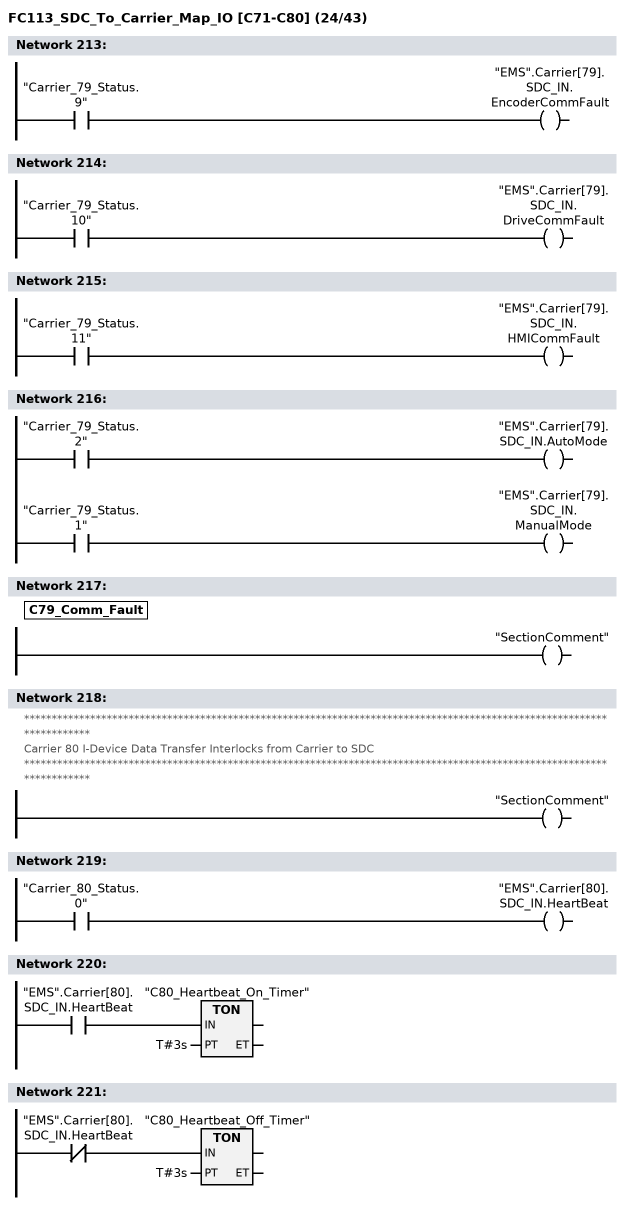
   RUNG wire#powerrail
      Contact( "Carrier_79_Status.9" )
      Coil( "EMS".Carrier[79].SDC_IN.EncoderCommFault )
   END_RUNG
   // the same network as SCL:
   "EMS".Carrier[79].SDC_IN.EncoderCommFault := "Carrier_79_Status.9";
END_REGION

REGION Network 214
   RUNG wire#powerrail
      Contact( "Carrier_79_Status.10" )
      Coil( "EMS".Carrier[79].SDC_IN.DriveCommFault )
   END_RUNG
   // the same network as SCL:
   "EMS".Carrier[79].SDC_IN.DriveCommFault := "Carrier_79_Status.10";
END_REGION

REGION Network 215
   RUNG wire#powerrail
      Contact( "Carrier_79_Status.11" )
      Coil( "EMS".Carrier[79].SDC_IN.HMICommFault )
   END_RUNG
   // the same network as SCL:
   "EMS".Carrier[79].SDC_IN.HMICommFault := "Carrier_79_Status.11";
END_REGION

REGION Network 216
   RUNG wire#powerrail
      Contact( "Carrier_79_Status.2" )
      Coil( "EMS".Carrier[79].SDC_IN.AutoMode )
   END_RUNG
   RUNG wire#powerrail
      Contact( "Carrier_79_Status.1" )
      Coil( "EMS".Carrier[79].SDC_IN.ManualMode )
   END_RUNG
   // the same network as SCL:
   "EMS".Carrier[79].SDC_IN.AutoMode := "Carrier_79_Status.2";
   "EMS".Carrier[79].SDC_IN.ManualMode := "Carrier_79_Status.1";
END_REGION

REGION Network 217
   Label( C79_Comm_Fault )
   RUNG wire#powerrail
      Coil( "SectionComment" )
   END_RUNG
   // the same network as SCL:
   C79_Comm_Fault:
   "SectionComment" := TRUE;
END_REGION

REGION Network 218
   // **********************************************************************************************************************
   // 
   // Carrier 80 I-Device Data Transfer Interlocks from Carrier to SDC
   // 
   // **********************************************************************************************************************
   RUNG wire#powerrail
      Coil( "SectionComment" )
   END_RUNG
   // the same network as SCL:
   "SectionComment" := TRUE;
END_REGION

REGION Network 219
   RUNG wire#powerrail
      Contact( "Carrier_80_Status.0" )
      Coil( "EMS".Carrier[80].SDC_IN.HeartBeat )
   END_RUNG
   // the same network as SCL:
   "EMS".Carrier[80].SDC_IN.HeartBeat := "Carrier_80_Status.0";
END_REGION

REGION Network 220
   "C80_Heartbeat_On_Timer".TON(IN := "EMS".Carrier[80].SDC_IN.HeartBeat, PT := T#3s);
END_REGION

REGION Network 221
   "C80_Heartbeat_Off_Timer".TON(IN := NOT "EMS".Carrier[80].SDC_IN.HeartBeat, PT := T#3s);
END_REGION

REGION Network 222
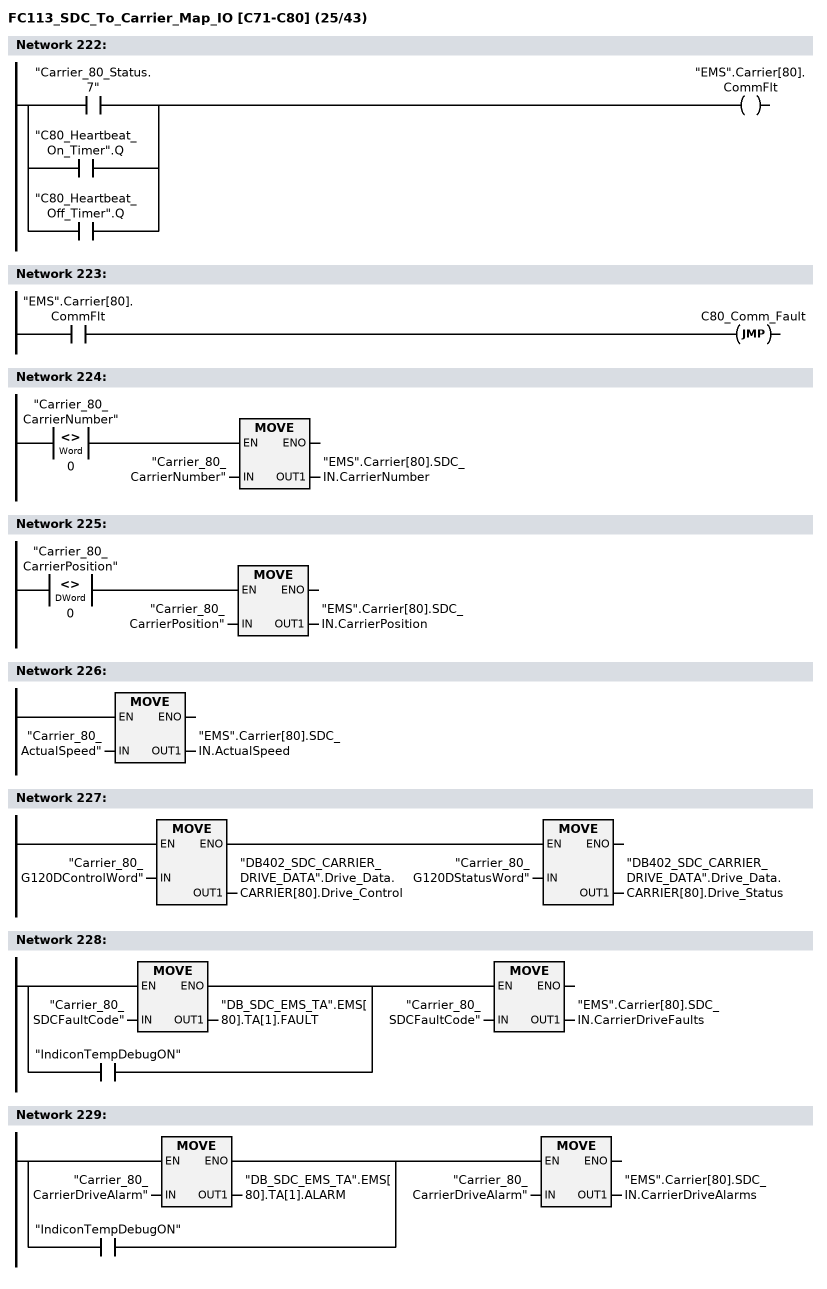
   RUNG wire#powerrail
      Contact( "Carrier_80_Status.7" )
      wire#w1
      Coil( "EMS".Carrier[80].CommFlt )
   END_RUNG
   RUNG wire#powerrail
      Contact( "C80_Heartbeat_On_Timer".Q )
   END_RUNG wire#w1
   RUNG wire#powerrail
      Contact( "C80_Heartbeat_Off_Timer".Q )
   END_RUNG wire#w1
   // the same network as SCL:
   "EMS".Carrier[80].CommFlt := "Carrier_80_Status.7" OR "C80_Heartbeat_On_Timer".Q OR "C80_Heartbeat_Off_Timer".Q;
END_REGION

REGION Network 223
   RUNG wire#powerrail
      Contact( "EMS".Carrier[80].CommFlt )
      JumpCoil( C80_Comm_Fault )
   END_RUNG
   // the same network as SCL:
   IF "EMS".Carrier[80].CommFlt THEN GOTO C80_Comm_Fault; END_IF;
END_REGION

REGION Network 224
   RUNG wire#powerrail
      { S7_Templates := "SrcType := Word" } NE_Contact(in1 := "Carrier_80_CarrierNumber", in2 := 0)
      Move(in := "Carrier_80_CarrierNumber", out1 => "EMS".Carrier[80].SDC_IN.CarrierNumber)
   END_RUNG
   // the same network as SCL:
   IF "Carrier_80_CarrierNumber" <> 0 THEN
       "EMS".Carrier[80].SDC_IN.CarrierNumber := "Carrier_80_CarrierNumber";
   END_IF;
END_REGION

REGION Network 225
   RUNG wire#powerrail
      { S7_Templates := "SrcType := DWord" } NE_Contact(in1 := "Carrier_80_CarrierPosition", in2 := 0)
      Move(in := "Carrier_80_CarrierPosition", out1 => "EMS".Carrier[80].SDC_IN.CarrierPosition)
   END_RUNG
   // the same network as SCL:
   IF "Carrier_80_CarrierPosition" <> 0 THEN
       "EMS".Carrier[80].SDC_IN.CarrierPosition := "Carrier_80_CarrierPosition";
   END_IF;
END_REGION

REGION Network 226
   RUNG wire#powerrail
      Move(in := "Carrier_80_ActualSpeed", out1 => "EMS".Carrier[80].SDC_IN.ActualSpeed)
   END_RUNG
   // the same network as SCL:
   "EMS".Carrier[80].SDC_IN.ActualSpeed := "Carrier_80_ActualSpeed";
END_REGION

REGION Network 227
   RUNG wire#powerrail
      Move(in := "Carrier_80_G120DControlWord", out1 => "DB402_SDC_CARRIER_DRIVE_DATA".Drive_Data.CARRIER[80].Drive_Control)
      Move(in := "Carrier_80_G120DStatusWord", out1 => "DB402_SDC_CARRIER_DRIVE_DATA".Drive_Data.CARRIER[80].Drive_Status)
   END_RUNG
   // the same network as SCL:
   "DB402_SDC_CARRIER_DRIVE_DATA".Drive_Data.CARRIER[80].Drive_Control := "Carrier_80_G120DControlWord";
   "DB402_SDC_CARRIER_DRIVE_DATA".Drive_Data.CARRIER[80].Drive_Status := "Carrier_80_G120DStatusWord";
END_REGION

REGION Network 228
   RUNG wire#powerrail
      Move(in := "Carrier_80_SDCFaultCode", out1 => "DB_SDC_EMS_TA".EMS[80].TA[1].FAULT)
      wire#w1
      Move(in := "Carrier_80_SDCFaultCode", out1 => "EMS".Carrier[80].SDC_IN.CarrierDriveFaults)
   END_RUNG
   RUNG wire#powerrail
      Contact( "IndiconTempDebugON" )
   END_RUNG wire#w1
   // the same network as SCL:
   "DB_SDC_EMS_TA".EMS[80].TA[1].FAULT := "Carrier_80_SDCFaultCode";
   IF TRUE OR "IndiconTempDebugON" THEN
       "EMS".Carrier[80].SDC_IN.CarrierDriveFaults := "Carrier_80_SDCFaultCode";
   END_IF;
END_REGION

REGION Network 229
   RUNG wire#powerrail
      Move(in := "Carrier_80_CarrierDriveAlarm", out1 => "DB_SDC_EMS_TA".EMS[80].TA[1].ALARM)
      wire#w1
      Move(in := "Carrier_80_CarrierDriveAlarm", out1 => "EMS".Carrier[80].SDC_IN.CarrierDriveAlarms)
   END_RUNG
   RUNG wire#powerrail
      Contact( "IndiconTempDebugON" )
   END_RUNG wire#w1
   // the same network as SCL:
   "DB_SDC_EMS_TA".EMS[80].TA[1].ALARM := "Carrier_80_CarrierDriveAlarm";
   IF TRUE OR "IndiconTempDebugON" THEN
       "EMS".Carrier[80].SDC_IN.CarrierDriveAlarms := "Carrier_80_CarrierDriveAlarm";
   END_IF;
END_REGION

REGION Network 230
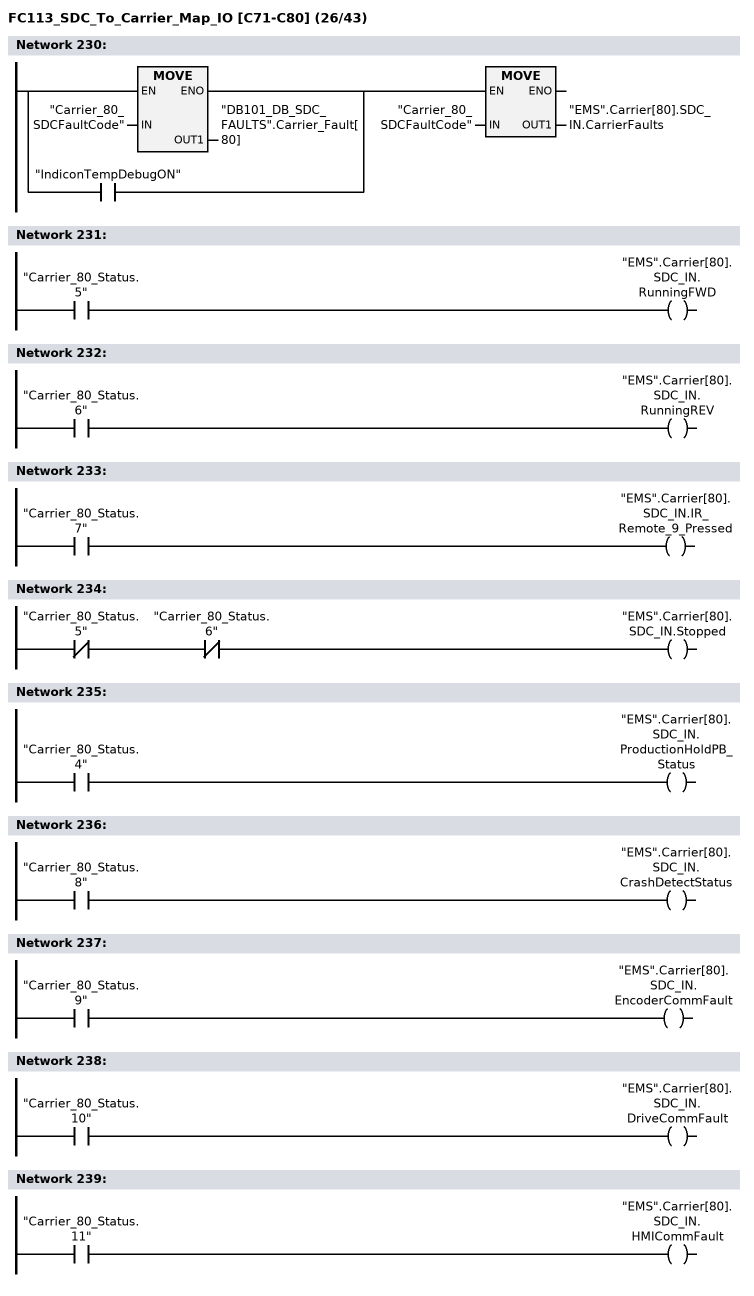
   RUNG wire#powerrail
      Move(in := "Carrier_80_SDCFaultCode", out1 => "DB101_DB_SDC_FAULTS".Carrier_Fault[80])
      wire#w1
      Move(in := "Carrier_80_SDCFaultCode", out1 => "EMS".Carrier[80].SDC_IN.CarrierFaults)
   END_RUNG
   RUNG wire#powerrail
      Contact( "IndiconTempDebugON" )
   END_RUNG wire#w1
   // the same network as SCL:
   "DB101_DB_SDC_FAULTS".Carrier_Fault[80] := "Carrier_80_SDCFaultCode";
   IF TRUE OR "IndiconTempDebugON" THEN
       "EMS".Carrier[80].SDC_IN.CarrierFaults := "Carrier_80_SDCFaultCode";
   END_IF;
END_REGION

REGION Network 231
   RUNG wire#powerrail
      Contact( "Carrier_80_Status.5" )
      Coil( "EMS".Carrier[80].SDC_IN.RunningFWD )
   END_RUNG
   // the same network as SCL:
   "EMS".Carrier[80].SDC_IN.RunningFWD := "Carrier_80_Status.5";
END_REGION

REGION Network 232
   RUNG wire#powerrail
      Contact( "Carrier_80_Status.6" )
      Coil( "EMS".Carrier[80].SDC_IN.RunningREV )
   END_RUNG
   // the same network as SCL:
   "EMS".Carrier[80].SDC_IN.RunningREV := "Carrier_80_Status.6";
END_REGION

REGION Network 233
   RUNG wire#powerrail
      Contact( "Carrier_80_Status.7" )
      Coil( "EMS".Carrier[80].SDC_IN.IR_Remote_9_Pressed )
   END_RUNG
   // the same network as SCL:
   "EMS".Carrier[80].SDC_IN.IR_Remote_9_Pressed := "Carrier_80_Status.7";
END_REGION

REGION Network 234
   RUNG wire#powerrail
      I_Contact( "Carrier_80_Status.5" )
      I_Contact( "Carrier_80_Status.6" )
      Coil( "EMS".Carrier[80].SDC_IN.Stopped )
   END_RUNG
   // the same network as SCL:
   "EMS".Carrier[80].SDC_IN.Stopped := NOT "Carrier_80_Status.5" AND NOT "Carrier_80_Status.6";
END_REGION

REGION Network 235
   RUNG wire#powerrail
      Contact( "Carrier_80_Status.4" )
      Coil( "EMS".Carrier[80].SDC_IN.ProductionHoldPB_Status )
   END_RUNG
   // the same network as SCL:
   "EMS".Carrier[80].SDC_IN.ProductionHoldPB_Status := "Carrier_80_Status.4";
END_REGION

REGION Network 236
   RUNG wire#powerrail
      Contact( "Carrier_80_Status.8" )
      Coil( "EMS".Carrier[80].SDC_IN.CrashDetectStatus )
   END_RUNG
   // the same network as SCL:
   "EMS".Carrier[80].SDC_IN.CrashDetectStatus := "Carrier_80_Status.8";
END_REGION

REGION Network 237
   RUNG wire#powerrail
      Contact( "Carrier_80_Status.9" )
      Coil( "EMS".Carrier[80].SDC_IN.EncoderCommFault )
   END_RUNG
   // the same network as SCL:
   "EMS".Carrier[80].SDC_IN.EncoderCommFault := "Carrier_80_Status.9";
END_REGION

REGION Network 238
   RUNG wire#powerrail
      Contact( "Carrier_80_Status.10" )
      Coil( "EMS".Carrier[80].SDC_IN.DriveCommFault )
   END_RUNG
   // the same network as SCL:
   "EMS".Carrier[80].SDC_IN.DriveCommFault := "Carrier_80_Status.10";
END_REGION

REGION Network 239
   RUNG wire#powerrail
      Contact( "Carrier_80_Status.11" )
      Coil( "EMS".Carrier[80].SDC_IN.HMICommFault )
   END_RUNG
   // the same network as SCL:
   "EMS".Carrier[80].SDC_IN.HMICommFault := "Carrier_80_Status.11";
END_REGION

REGION Network 240
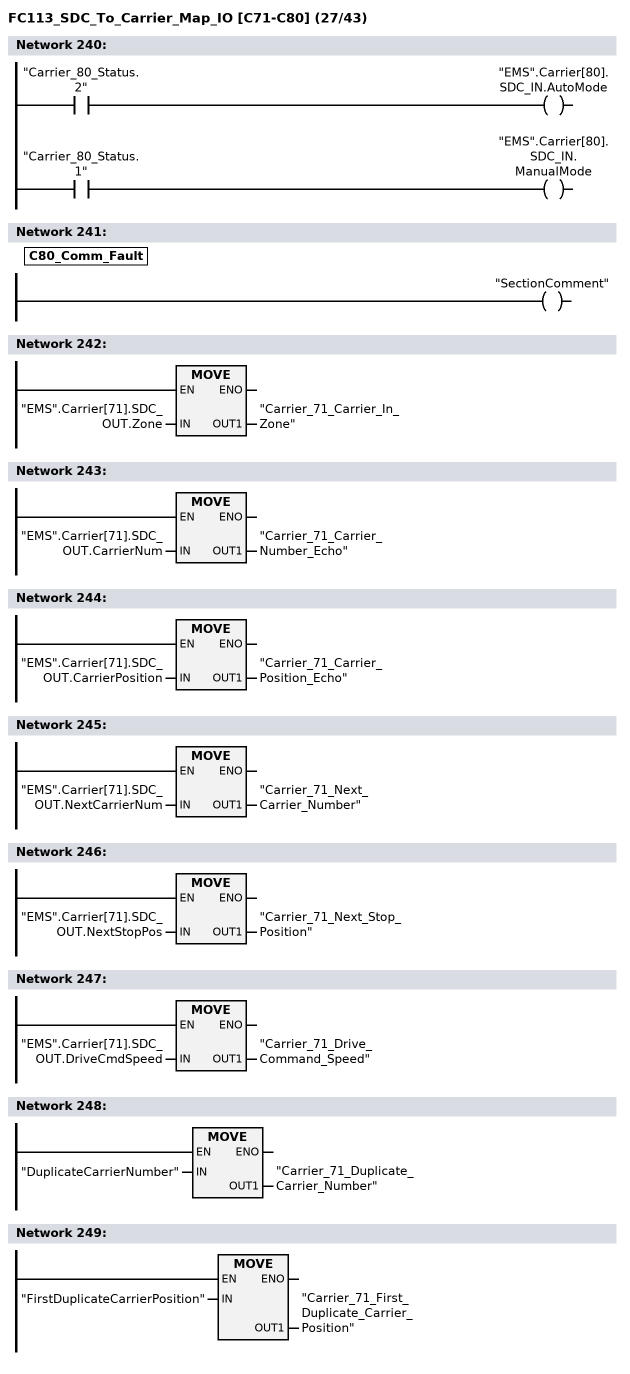
   RUNG wire#powerrail
      Contact( "Carrier_80_Status.2" )
      Coil( "EMS".Carrier[80].SDC_IN.AutoMode )
   END_RUNG
   RUNG wire#powerrail
      Contact( "Carrier_80_Status.1" )
      Coil( "EMS".Carrier[80].SDC_IN.ManualMode )
   END_RUNG
   // the same network as SCL:
   "EMS".Carrier[80].SDC_IN.AutoMode := "Carrier_80_Status.2";
   "EMS".Carrier[80].SDC_IN.ManualMode := "Carrier_80_Status.1";
END_REGION

REGION Network 241
   Label( C80_Comm_Fault )
   RUNG wire#powerrail
      Coil( "SectionComment" )
   END_RUNG
   // the same network as SCL:
   C80_Comm_Fault:
   "SectionComment" := TRUE;
END_REGION

REGION Network 242
   RUNG wire#powerrail
      Move(in := "EMS".Carrier[71].SDC_OUT.Zone, out1 => "Carrier_71_Carrier_In_Zone")
   END_RUNG
   // the same network as SCL:
   "Carrier_71_Carrier_In_Zone" := "EMS".Carrier[71].SDC_OUT.Zone;
END_REGION

REGION Network 243
   RUNG wire#powerrail
      Move(in := "EMS".Carrier[71].SDC_OUT.CarrierNum, out1 => "Carrier_71_Carrier_Number_Echo")
   END_RUNG
   // the same network as SCL:
   "Carrier_71_Carrier_Number_Echo" := "EMS".Carrier[71].SDC_OUT.CarrierNum;
END_REGION

REGION Network 244
   RUNG wire#powerrail
      Move(in := "EMS".Carrier[71].SDC_OUT.CarrierPosition, out1 => "Carrier_71_Carrier_Position_Echo")
   END_RUNG
   // the same network as SCL:
   "Carrier_71_Carrier_Position_Echo" := "EMS".Carrier[71].SDC_OUT.CarrierPosition;
END_REGION

REGION Network 245
   RUNG wire#powerrail
      Move(in := "EMS".Carrier[71].SDC_OUT.NextCarrierNum, out1 => "Carrier_71_Next_Carrier_Number")
   END_RUNG
   // the same network as SCL:
   "Carrier_71_Next_Carrier_Number" := "EMS".Carrier[71].SDC_OUT.NextCarrierNum;
END_REGION

REGION Network 246
   RUNG wire#powerrail
      Move(in := "EMS".Carrier[71].SDC_OUT.NextStopPos, out1 => "Carrier_71_Next_Stop_Position")
   END_RUNG
   // the same network as SCL:
   "Carrier_71_Next_Stop_Position" := "EMS".Carrier[71].SDC_OUT.NextStopPos;
END_REGION

REGION Network 247
   RUNG wire#powerrail
      Move(in := "EMS".Carrier[71].SDC_OUT.DriveCmdSpeed, out1 => "Carrier_71_Drive_Command_Speed")
   END_RUNG
   // the same network as SCL:
   "Carrier_71_Drive_Command_Speed" := "EMS".Carrier[71].SDC_OUT.DriveCmdSpeed;
END_REGION

REGION Network 248
   RUNG wire#powerrail
      Move(in := "DuplicateCarrierNumber", out1 => "Carrier_71_Duplicate_Carrier_Number")
   END_RUNG
   // the same network as SCL:
   "Carrier_71_Duplicate_Carrier_Number" := "DuplicateCarrierNumber";
END_REGION

REGION Network 249
   RUNG wire#powerrail
      Move(in := "FirstDuplicateCarrierPosition", out1 => "Carrier_71_First_Duplicate_Carrier_Position")
   END_RUNG
   // the same network as SCL:
   "Carrier_71_First_Duplicate_Carrier_Position" := "FirstDuplicateCarrierPosition";
END_REGION

REGION Network 250
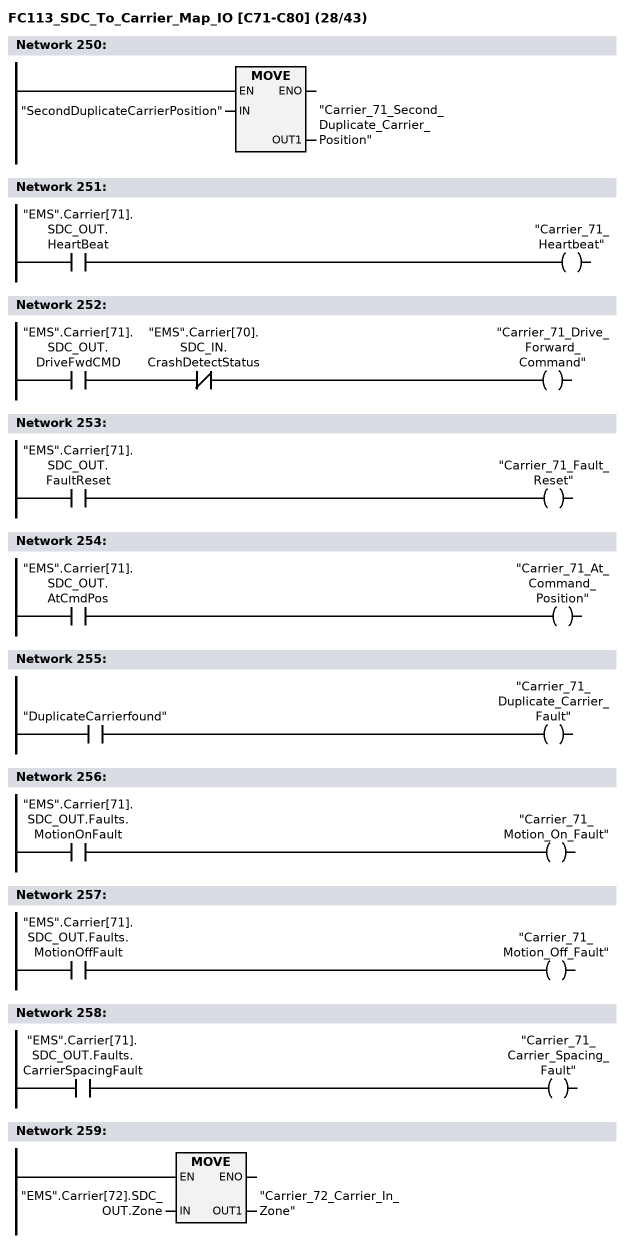
   RUNG wire#powerrail
      Move(in := "SecondDuplicateCarrierPosition", out1 => "Carrier_71_Second_Duplicate_Carrier_Position")
   END_RUNG
   // the same network as SCL:
   "Carrier_71_Second_Duplicate_Carrier_Position" := "SecondDuplicateCarrierPosition";
END_REGION

REGION Network 251
   RUNG wire#powerrail
      Contact( "EMS".Carrier[71].SDC_OUT.HeartBeat )
      Coil( "Carrier_71_Heartbeat" )
   END_RUNG
   // the same network as SCL:
   "Carrier_71_Heartbeat" := "EMS".Carrier[71].SDC_OUT.HeartBeat;
END_REGION

REGION Network 252
   RUNG wire#powerrail
      Contact( "EMS".Carrier[71].SDC_OUT.DriveFwdCMD )
      I_Contact( "EMS".Carrier[70].SDC_IN.CrashDetectStatus )
      Coil( "Carrier_71_Drive_Forward_Command" )
   END_RUNG
   // the same network as SCL:
   "Carrier_71_Drive_Forward_Command" := "EMS".Carrier[71].SDC_OUT.DriveFwdCMD AND NOT "EMS".Carrier[70].SDC_IN.CrashDetectStatus;
END_REGION

REGION Network 253
   RUNG wire#powerrail
      Contact( "EMS".Carrier[71].SDC_OUT.FaultReset )
      Coil( "Carrier_71_Fault_Reset" )
   END_RUNG
   // the same network as SCL:
   "Carrier_71_Fault_Reset" := "EMS".Carrier[71].SDC_OUT.FaultReset;
END_REGION

REGION Network 254
   RUNG wire#powerrail
      Contact( "EMS".Carrier[71].SDC_OUT.AtCmdPos )
      Coil( "Carrier_71_At_Command_Position" )
   END_RUNG
   // the same network as SCL:
   "Carrier_71_At_Command_Position" := "EMS".Carrier[71].SDC_OUT.AtCmdPos;
END_REGION

REGION Network 255
   RUNG wire#powerrail
      Contact( "DuplicateCarrierfound" )
      Coil( "Carrier_71_Duplicate_Carrier_Fault" )
   END_RUNG
   // the same network as SCL:
   "Carrier_71_Duplicate_Carrier_Fault" := "DuplicateCarrierfound";
END_REGION

REGION Network 256
   RUNG wire#powerrail
      Contact( "EMS".Carrier[71].SDC_OUT.Faults.MotionOnFault )
      Coil( "Carrier_71_Motion_On_Fault" )
   END_RUNG
   // the same network as SCL:
   "Carrier_71_Motion_On_Fault" := "EMS".Carrier[71].SDC_OUT.Faults.MotionOnFault;
END_REGION

REGION Network 257
   RUNG wire#powerrail
      Contact( "EMS".Carrier[71].SDC_OUT.Faults.MotionOffFault )
      Coil( "Carrier_71_Motion_Off_Fault" )
   END_RUNG
   // the same network as SCL:
   "Carrier_71_Motion_Off_Fault" := "EMS".Carrier[71].SDC_OUT.Faults.MotionOffFault;
END_REGION

REGION Network 258
   RUNG wire#powerrail
      Contact( "EMS".Carrier[71].SDC_OUT.Faults.CarrierSpacingFault )
      Coil( "Carrier_71_Carrier_Spacing_Fault" )
   END_RUNG
   // the same network as SCL:
   "Carrier_71_Carrier_Spacing_Fault" := "EMS".Carrier[71].SDC_OUT.Faults.CarrierSpacingFault;
END_REGION

REGION Network 259
   RUNG wire#powerrail
      Move(in := "EMS".Carrier[72].SDC_OUT.Zone, out1 => "Carrier_72_Carrier_In_Zone")
   END_RUNG
   // the same network as SCL:
   "Carrier_72_Carrier_In_Zone" := "EMS".Carrier[72].SDC_OUT.Zone;
END_REGION

REGION Network 260
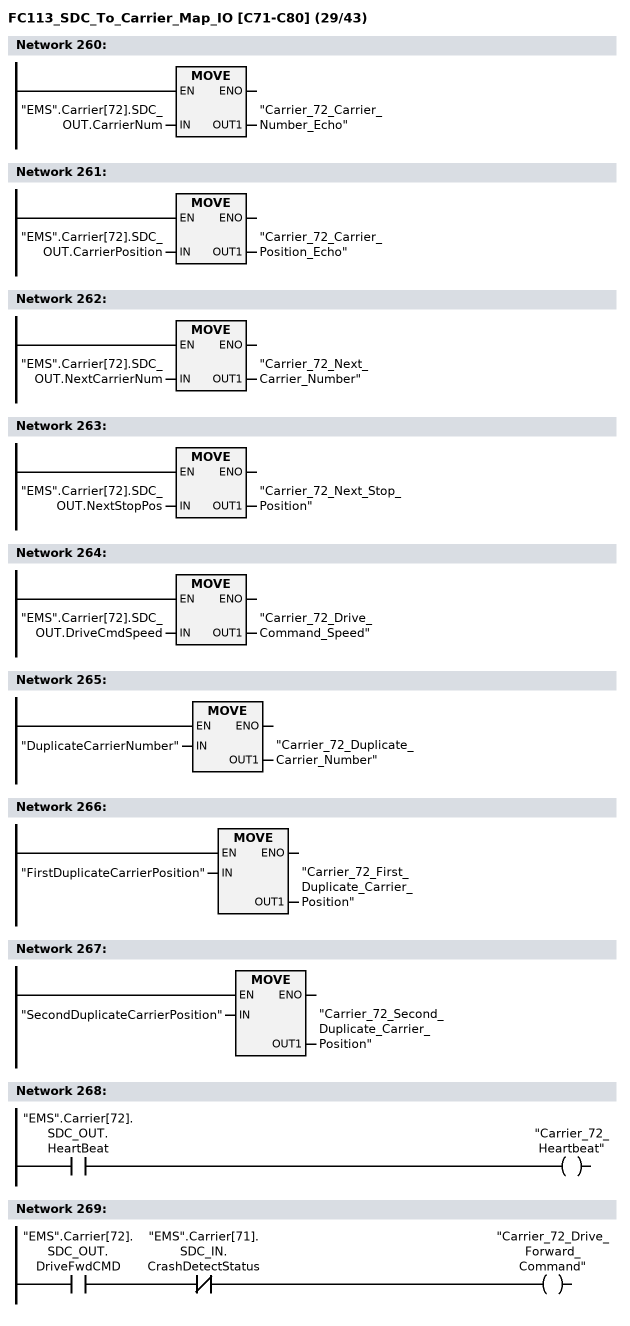
   RUNG wire#powerrail
      Move(in := "EMS".Carrier[72].SDC_OUT.CarrierNum, out1 => "Carrier_72_Carrier_Number_Echo")
   END_RUNG
   // the same network as SCL:
   "Carrier_72_Carrier_Number_Echo" := "EMS".Carrier[72].SDC_OUT.CarrierNum;
END_REGION

REGION Network 261
   RUNG wire#powerrail
      Move(in := "EMS".Carrier[72].SDC_OUT.CarrierPosition, out1 => "Carrier_72_Carrier_Position_Echo")
   END_RUNG
   // the same network as SCL:
   "Carrier_72_Carrier_Position_Echo" := "EMS".Carrier[72].SDC_OUT.CarrierPosition;
END_REGION

REGION Network 262
   RUNG wire#powerrail
      Move(in := "EMS".Carrier[72].SDC_OUT.NextCarrierNum, out1 => "Carrier_72_Next_Carrier_Number")
   END_RUNG
   // the same network as SCL:
   "Carrier_72_Next_Carrier_Number" := "EMS".Carrier[72].SDC_OUT.NextCarrierNum;
END_REGION

REGION Network 263
   RUNG wire#powerrail
      Move(in := "EMS".Carrier[72].SDC_OUT.NextStopPos, out1 => "Carrier_72_Next_Stop_Position")
   END_RUNG
   // the same network as SCL:
   "Carrier_72_Next_Stop_Position" := "EMS".Carrier[72].SDC_OUT.NextStopPos;
END_REGION

REGION Network 264
   RUNG wire#powerrail
      Move(in := "EMS".Carrier[72].SDC_OUT.DriveCmdSpeed, out1 => "Carrier_72_Drive_Command_Speed")
   END_RUNG
   // the same network as SCL:
   "Carrier_72_Drive_Command_Speed" := "EMS".Carrier[72].SDC_OUT.DriveCmdSpeed;
END_REGION

REGION Network 265
   RUNG wire#powerrail
      Move(in := "DuplicateCarrierNumber", out1 => "Carrier_72_Duplicate_Carrier_Number")
   END_RUNG
   // the same network as SCL:
   "Carrier_72_Duplicate_Carrier_Number" := "DuplicateCarrierNumber";
END_REGION

REGION Network 266
   RUNG wire#powerrail
      Move(in := "FirstDuplicateCarrierPosition", out1 => "Carrier_72_First_Duplicate_Carrier_Position")
   END_RUNG
   // the same network as SCL:
   "Carrier_72_First_Duplicate_Carrier_Position" := "FirstDuplicateCarrierPosition";
END_REGION

REGION Network 267
   RUNG wire#powerrail
      Move(in := "SecondDuplicateCarrierPosition", out1 => "Carrier_72_Second_Duplicate_Carrier_Position")
   END_RUNG
   // the same network as SCL:
   "Carrier_72_Second_Duplicate_Carrier_Position" := "SecondDuplicateCarrierPosition";
END_REGION

REGION Network 268
   RUNG wire#powerrail
      Contact( "EMS".Carrier[72].SDC_OUT.HeartBeat )
      Coil( "Carrier_72_Heartbeat" )
   END_RUNG
   // the same network as SCL:
   "Carrier_72_Heartbeat" := "EMS".Carrier[72].SDC_OUT.HeartBeat;
END_REGION

REGION Network 269
   RUNG wire#powerrail
      Contact( "EMS".Carrier[72].SDC_OUT.DriveFwdCMD )
      I_Contact( "EMS".Carrier[71].SDC_IN.CrashDetectStatus )
      Coil( "Carrier_72_Drive_Forward_Command" )
   END_RUNG
   // the same network as SCL:
   "Carrier_72_Drive_Forward_Command" := "EMS".Carrier[72].SDC_OUT.DriveFwdCMD AND NOT "EMS".Carrier[71].SDC_IN.CrashDetectStatus;
END_REGION

REGION Network 270
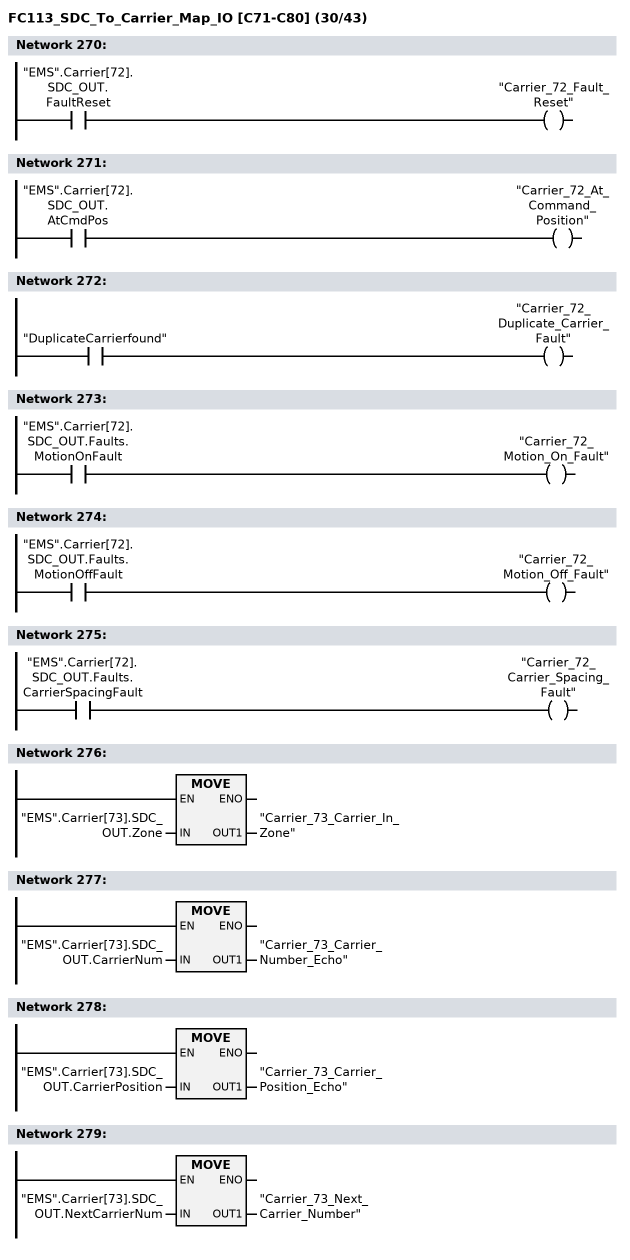
   RUNG wire#powerrail
      Contact( "EMS".Carrier[72].SDC_OUT.FaultReset )
      Coil( "Carrier_72_Fault_Reset" )
   END_RUNG
   // the same network as SCL:
   "Carrier_72_Fault_Reset" := "EMS".Carrier[72].SDC_OUT.FaultReset;
END_REGION

REGION Network 271
   RUNG wire#powerrail
      Contact( "EMS".Carrier[72].SDC_OUT.AtCmdPos )
      Coil( "Carrier_72_At_Command_Position" )
   END_RUNG
   // the same network as SCL:
   "Carrier_72_At_Command_Position" := "EMS".Carrier[72].SDC_OUT.AtCmdPos;
END_REGION

REGION Network 272
   RUNG wire#powerrail
      Contact( "DuplicateCarrierfound" )
      Coil( "Carrier_72_Duplicate_Carrier_Fault" )
   END_RUNG
   // the same network as SCL:
   "Carrier_72_Duplicate_Carrier_Fault" := "DuplicateCarrierfound";
END_REGION

REGION Network 273
   RUNG wire#powerrail
      Contact( "EMS".Carrier[72].SDC_OUT.Faults.MotionOnFault )
      Coil( "Carrier_72_Motion_On_Fault" )
   END_RUNG
   // the same network as SCL:
   "Carrier_72_Motion_On_Fault" := "EMS".Carrier[72].SDC_OUT.Faults.MotionOnFault;
END_REGION

REGION Network 274
   RUNG wire#powerrail
      Contact( "EMS".Carrier[72].SDC_OUT.Faults.MotionOffFault )
      Coil( "Carrier_72_Motion_Off_Fault" )
   END_RUNG
   // the same network as SCL:
   "Carrier_72_Motion_Off_Fault" := "EMS".Carrier[72].SDC_OUT.Faults.MotionOffFault;
END_REGION

REGION Network 275
   RUNG wire#powerrail
      Contact( "EMS".Carrier[72].SDC_OUT.Faults.CarrierSpacingFault )
      Coil( "Carrier_72_Carrier_Spacing_Fault" )
   END_RUNG
   // the same network as SCL:
   "Carrier_72_Carrier_Spacing_Fault" := "EMS".Carrier[72].SDC_OUT.Faults.CarrierSpacingFault;
END_REGION

REGION Network 276
   RUNG wire#powerrail
      Move(in := "EMS".Carrier[73].SDC_OUT.Zone, out1 => "Carrier_73_Carrier_In_Zone")
   END_RUNG
   // the same network as SCL:
   "Carrier_73_Carrier_In_Zone" := "EMS".Carrier[73].SDC_OUT.Zone;
END_REGION

REGION Network 277
   RUNG wire#powerrail
      Move(in := "EMS".Carrier[73].SDC_OUT.CarrierNum, out1 => "Carrier_73_Carrier_Number_Echo")
   END_RUNG
   // the same network as SCL:
   "Carrier_73_Carrier_Number_Echo" := "EMS".Carrier[73].SDC_OUT.CarrierNum;
END_REGION

REGION Network 278
   RUNG wire#powerrail
      Move(in := "EMS".Carrier[73].SDC_OUT.CarrierPosition, out1 => "Carrier_73_Carrier_Position_Echo")
   END_RUNG
   // the same network as SCL:
   "Carrier_73_Carrier_Position_Echo" := "EMS".Carrier[73].SDC_OUT.CarrierPosition;
END_REGION

REGION Network 279
   RUNG wire#powerrail
      Move(in := "EMS".Carrier[73].SDC_OUT.NextCarrierNum, out1 => "Carrier_73_Next_Carrier_Number")
   END_RUNG
   // the same network as SCL:
   "Carrier_73_Next_Carrier_Number" := "EMS".Carrier[73].SDC_OUT.NextCarrierNum;
END_REGION

REGION Network 280
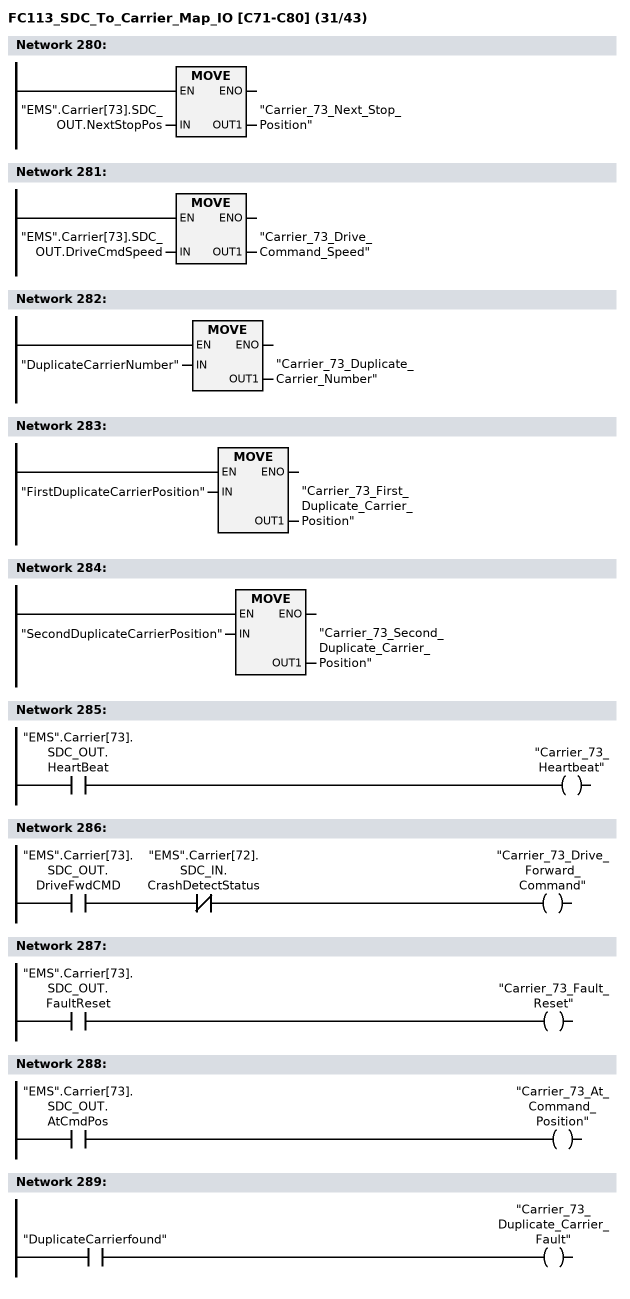
   RUNG wire#powerrail
      Move(in := "EMS".Carrier[73].SDC_OUT.NextStopPos, out1 => "Carrier_73_Next_Stop_Position")
   END_RUNG
   // the same network as SCL:
   "Carrier_73_Next_Stop_Position" := "EMS".Carrier[73].SDC_OUT.NextStopPos;
END_REGION

REGION Network 281
   RUNG wire#powerrail
      Move(in := "EMS".Carrier[73].SDC_OUT.DriveCmdSpeed, out1 => "Carrier_73_Drive_Command_Speed")
   END_RUNG
   // the same network as SCL:
   "Carrier_73_Drive_Command_Speed" := "EMS".Carrier[73].SDC_OUT.DriveCmdSpeed;
END_REGION

REGION Network 282
   RUNG wire#powerrail
      Move(in := "DuplicateCarrierNumber", out1 => "Carrier_73_Duplicate_Carrier_Number")
   END_RUNG
   // the same network as SCL:
   "Carrier_73_Duplicate_Carrier_Number" := "DuplicateCarrierNumber";
END_REGION

REGION Network 283
   RUNG wire#powerrail
      Move(in := "FirstDuplicateCarrierPosition", out1 => "Carrier_73_First_Duplicate_Carrier_Position")
   END_RUNG
   // the same network as SCL:
   "Carrier_73_First_Duplicate_Carrier_Position" := "FirstDuplicateCarrierPosition";
END_REGION

REGION Network 284
   RUNG wire#powerrail
      Move(in := "SecondDuplicateCarrierPosition", out1 => "Carrier_73_Second_Duplicate_Carrier_Position")
   END_RUNG
   // the same network as SCL:
   "Carrier_73_Second_Duplicate_Carrier_Position" := "SecondDuplicateCarrierPosition";
END_REGION

REGION Network 285
   RUNG wire#powerrail
      Contact( "EMS".Carrier[73].SDC_OUT.HeartBeat )
      Coil( "Carrier_73_Heartbeat" )
   END_RUNG
   // the same network as SCL:
   "Carrier_73_Heartbeat" := "EMS".Carrier[73].SDC_OUT.HeartBeat;
END_REGION

REGION Network 286
   RUNG wire#powerrail
      Contact( "EMS".Carrier[73].SDC_OUT.DriveFwdCMD )
      I_Contact( "EMS".Carrier[72].SDC_IN.CrashDetectStatus )
      Coil( "Carrier_73_Drive_Forward_Command" )
   END_RUNG
   // the same network as SCL:
   "Carrier_73_Drive_Forward_Command" := "EMS".Carrier[73].SDC_OUT.DriveFwdCMD AND NOT "EMS".Carrier[72].SDC_IN.CrashDetectStatus;
END_REGION

REGION Network 287
   RUNG wire#powerrail
      Contact( "EMS".Carrier[73].SDC_OUT.FaultReset )
      Coil( "Carrier_73_Fault_Reset" )
   END_RUNG
   // the same network as SCL:
   "Carrier_73_Fault_Reset" := "EMS".Carrier[73].SDC_OUT.FaultReset;
END_REGION

REGION Network 288
   RUNG wire#powerrail
      Contact( "EMS".Carrier[73].SDC_OUT.AtCmdPos )
      Coil( "Carrier_73_At_Command_Position" )
   END_RUNG
   // the same network as SCL:
   "Carrier_73_At_Command_Position" := "EMS".Carrier[73].SDC_OUT.AtCmdPos;
END_REGION

REGION Network 289
   RUNG wire#powerrail
      Contact( "DuplicateCarrierfound" )
      Coil( "Carrier_73_Duplicate_Carrier_Fault" )
   END_RUNG
   // the same network as SCL:
   "Carrier_73_Duplicate_Carrier_Fault" := "DuplicateCarrierfound";
END_REGION

REGION Network 290
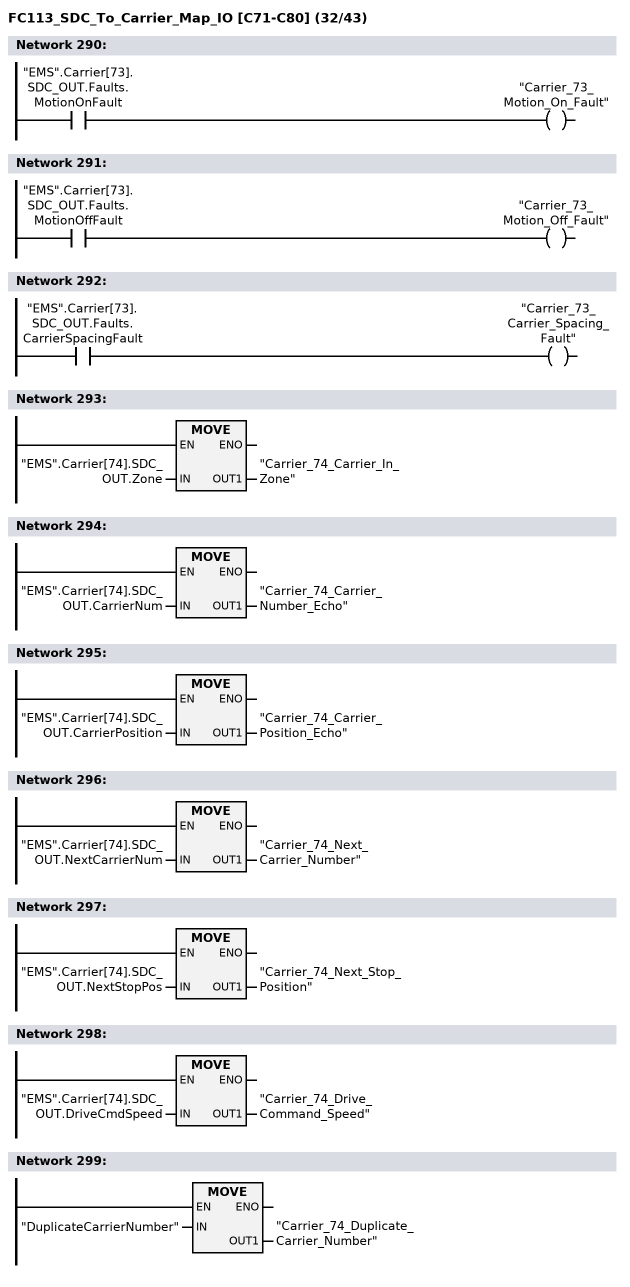
   RUNG wire#powerrail
      Contact( "EMS".Carrier[73].SDC_OUT.Faults.MotionOnFault )
      Coil( "Carrier_73_Motion_On_Fault" )
   END_RUNG
   // the same network as SCL:
   "Carrier_73_Motion_On_Fault" := "EMS".Carrier[73].SDC_OUT.Faults.MotionOnFault;
END_REGION

REGION Network 291
   RUNG wire#powerrail
      Contact( "EMS".Carrier[73].SDC_OUT.Faults.MotionOffFault )
      Coil( "Carrier_73_Motion_Off_Fault" )
   END_RUNG
   // the same network as SCL:
   "Carrier_73_Motion_Off_Fault" := "EMS".Carrier[73].SDC_OUT.Faults.MotionOffFault;
END_REGION

REGION Network 292
   RUNG wire#powerrail
      Contact( "EMS".Carrier[73].SDC_OUT.Faults.CarrierSpacingFault )
      Coil( "Carrier_73_Carrier_Spacing_Fault" )
   END_RUNG
   // the same network as SCL:
   "Carrier_73_Carrier_Spacing_Fault" := "EMS".Carrier[73].SDC_OUT.Faults.CarrierSpacingFault;
END_REGION

REGION Network 293
   RUNG wire#powerrail
      Move(in := "EMS".Carrier[74].SDC_OUT.Zone, out1 => "Carrier_74_Carrier_In_Zone")
   END_RUNG
   // the same network as SCL:
   "Carrier_74_Carrier_In_Zone" := "EMS".Carrier[74].SDC_OUT.Zone;
END_REGION

REGION Network 294
   RUNG wire#powerrail
      Move(in := "EMS".Carrier[74].SDC_OUT.CarrierNum, out1 => "Carrier_74_Carrier_Number_Echo")
   END_RUNG
   // the same network as SCL:
   "Carrier_74_Carrier_Number_Echo" := "EMS".Carrier[74].SDC_OUT.CarrierNum;
END_REGION

REGION Network 295
   RUNG wire#powerrail
      Move(in := "EMS".Carrier[74].SDC_OUT.CarrierPosition, out1 => "Carrier_74_Carrier_Position_Echo")
   END_RUNG
   // the same network as SCL:
   "Carrier_74_Carrier_Position_Echo" := "EMS".Carrier[74].SDC_OUT.CarrierPosition;
END_REGION

REGION Network 296
   RUNG wire#powerrail
      Move(in := "EMS".Carrier[74].SDC_OUT.NextCarrierNum, out1 => "Carrier_74_Next_Carrier_Number")
   END_RUNG
   // the same network as SCL:
   "Carrier_74_Next_Carrier_Number" := "EMS".Carrier[74].SDC_OUT.NextCarrierNum;
END_REGION

REGION Network 297
   RUNG wire#powerrail
      Move(in := "EMS".Carrier[74].SDC_OUT.NextStopPos, out1 => "Carrier_74_Next_Stop_Position")
   END_RUNG
   // the same network as SCL:
   "Carrier_74_Next_Stop_Position" := "EMS".Carrier[74].SDC_OUT.NextStopPos;
END_REGION

REGION Network 298
   RUNG wire#powerrail
      Move(in := "EMS".Carrier[74].SDC_OUT.DriveCmdSpeed, out1 => "Carrier_74_Drive_Command_Speed")
   END_RUNG
   // the same network as SCL:
   "Carrier_74_Drive_Command_Speed" := "EMS".Carrier[74].SDC_OUT.DriveCmdSpeed;
END_REGION

REGION Network 299
   RUNG wire#powerrail
      Move(in := "DuplicateCarrierNumber", out1 => "Carrier_74_Duplicate_Carrier_Number")
   END_RUNG
   // the same network as SCL:
   "Carrier_74_Duplicate_Carrier_Number" := "DuplicateCarrierNumber";
END_REGION

REGION Network 300
